
                   //Inner gross glass width [mm]
                   Chars_TO_Strg(Chars:=#AUX_rgcReceiveBuffer,
                                 pChars:=38,
                                 Cnt:=5,
                                 Strg=>#TMP_strValue);

                   #AUX_tYTelegram.dInLimitGross_mm := STRING_TO_DINT(#TMP_strValue); 

                   //Outer gross glass width [mm]
                   Chars_TO_Strg(Chars:=#AUX_rgcReceiveBuffer,
                                 pChars:=44,
                                 Cnt:=5,
                                 Strg=>#TMP_strValue);

                   #AUX_tYTelegram.dOutLimitGross_mm := STRING_TO_DINT(#TMP_strValue); 

                   //Center orientated position of the inner toproller [mm]
                   Chars_TO_Strg(Chars:=#AUX_rgcReceiveBuffer,
                                 pChars:=50,
                                 Cnt:=5,
                                 Strg=>#TMP_strValue);

                   #AUX_tYTelegram.dCenterOrientInTop_mm := STRING_TO_DINT(#TMP_strValue); 

                   //Edge orientated position of the inner toproller [mm]
                   Chars_TO_Strg(Chars:=#AUX_rgcReceiveBuffer,
                                 pChars:=56,
                                 Cnt:=5,
                                 Strg=>#TMP_strValue);

                   #AUX_tYTelegram.dEdgeOrientInTop_mm := STRING_TO_DINT(#TMP_strValue); 

                   //Center orientated position of the outer toproller [mm]
                   Chars_TO_Strg(Chars:=#AUX_rgcReceiveBuffer,
                                 pChars:=62,
                                 Cnt:=5,
                                 Strg=>#TMP_strValue);

                   #AUX_tYTelegram.dCenterOrientOutTop_mm := STRING_TO_DINT(#TMP_strValue); 

                   //Edge orientated position of the outer toproll [mm]
                   Chars_TO_Strg(Chars:=#AUX_rgcReceiveBuffer,
                                 pChars:=68,
                                 Cnt:=5,
                                 Strg=>#TMP_strValue);

                   #AUX_tYTelegram.dEdgeOrientOutTop_mm := STRING_TO_DINT(#TMP_strValue); 

                   //Check the conformity
                   IF #AUX_tYTelegram.dTelCounter < 0 OR
                      #AUX_tYTelegram.dTelCounter > 65535 OR
                      #AUX_tYTelegram.dFeedPulse_mm < 0 OR 
                      #AUX_tYTelegram.dFeedPulse_mm > 65535 OR
                      #AUX_tYTelegram.dInLimit_mm < 0 OR 
                      #AUX_tYTelegram.dInLimit_mm > 65535 OR
                      #AUX_tYTelegram.dOutLimit_mm < 0 OR 
                      #AUX_tYTelegram.dOutLimit_mm > 65535 OR
                      #AUX_tYTelegram.dInLimitUsable_mm < 0 OR 
                      #AUX_tYTelegram.dInLimitUsable_mm > 65535 OR
                      #AUX_tYTelegram.dOutLimitUsable_mm < 0 OR 
                      #AUX_tYTelegram.dOutLimitUsable_mm > 65535 OR
                      #AUX_tYTelegram.dInLimitGross_mm < 0 OR 
                      #AUX_tYTelegram.dInLimitGross_mm > 65535 OR
                      #AUX_tYTelegram.dOutLimitGross_mm < 0 OR 
                      #AUX_tYTelegram.dOutLimitGross_mm > 65535 OR
                      #AUX_tYTelegram.dCenterOrientInTop_mm < 0 OR 
                      #AUX_tYTelegram.dCenterOrientInTop_mm > 65535 OR
                      #AUX_tYTelegram.dEdgeOrientInTop_mm < 0 OR 
                      #AUX_tYTelegram.dEdgeOrientInTop_mm > 65535 OR
                      #AUX_tYTelegram.dCenterOrientOutTop_mm < 0 OR 
                      #AUX_tYTelegram.dCenterOrientOutTop_mm > 65535 OR
                      #AUX_tYTelegram.dEdgeOrientOutTop_mm < 0 OR 
                      #AUX_tYTelegram.dEdgeOrientOutTop_mm > 65535 THEN
                       #AUX_xTelegramYError := TRUE;
                   ELSE
                       IF #ST_xMachineSyncronized AND #tHMW.xAutoInspEnabled THEN

                           #TMP_dCountPos_cmm := #AUX_tYTelegram.dFeedPulse_mm - #AUX_dISRAValidCountMeter_mm;

                           IF #TMP_dCountPos_cmm < -32767 THEN

                               #AUX_tYTelegram.dPLCPosCount_cmm  := #AUX_dPLCValidCountMeter_cmm + ((#TMP_dCountPos_cmm + 65536)*100);

                           ELSIF #TMP_dCountPos_cmm > 32767 THEN

                               #AUX_tYTelegram.dPLCPosCount_cmm := #AUX_dPLCValidCountMeter_cmm + ((#TMP_dCountPos_cmm - 65536)*100);

                           ELSE

                               #AUX_tYTelegram.dPLCPosCount_cmm := #AUX_dPLCValidCountMeter_cmm + (#TMP_dCountPos_cmm * 100);

                           END_IF;

                           #AUX_tYTelegram.dPLCPosCount_cmm := #tHMR.dDistSnapRoll_cmm + #AUX_tYTelegram.dPLCPosCount_cmm;

                           #tHMR.dCurrentGrossWidth_cmm := (#AUX_tYTelegram.dOutLimitGross_mm - #AUX_tYTelegram.dInLimitGross_mm) * 100 ;
                           #tHMR.dCurrentNetWidth_cmm := (#AUX_tYTelegram.dOutLimitUsable_mm - #AUX_tYTelegram.dInLimitUsable_mm) * 100 ;

                           IF (#tHMR.dDistCenterLine_cmm <= 0) THEN

                               #tHMR.dCurrentGrossWander_cmm := #tHMR.dDistCenterLine_cmm + ((#AUX_tYTelegram.dInLimitGross_mm + #AUX_tYTelegram.dOutLimitGross_mm)/2) * 100;
                               #tHMR.dCurrentNetWander_cmm := #tHMR.dDistCenterLine_cmm + ((#AUX_tYTelegram.dInLimitUsable_mm + #AUX_tYTelegram.dOutLimitUsable_mm)/2) * 100;

                           ELSE
                               #tHMR.dCurrentGrossWander_cmm := #tHMR.dDistCenterLine_cmm - ((#AUX_tYTelegram.dInLimitGross_mm + #AUX_tYTelegram.dOutLimitGross_mm)/2) * 100;
                               #tHMR.dCurrentNetWander_cmm := #tHMR.dDistCenterLine_cmm - ((#AUX_tYTelegram.dInLimitUsable_mm + #AUX_tYTelegram.dOutLimitUsable_mm)/2) * 100;

                           END_IF;

                           #INO_tRibbon.rgtGlassData[#IN_dGlassDataMachineIndex].dDistSnapRoll_cmm := #tHMR.dDistSnapRoll_cmm + #DISRADEADPOINT_CMM; 

                           //Update the position
                           IF NOT #INO_tRibbon.rgtGlassDataUpdate[#IN_dGlassDataUpdateMachineIndex].xUpdateRequest THEN
                               #INO_tRibbon.rgtGlassDataUpdate[#IN_dGlassDataUpdateMachineIndex].tData.dGrossWander_cmm := #tHMR.dCurrentGrossWander_cmm;
                               #INO_tRibbon.rgtGlassDataUpdate[#IN_dGlassDataUpdateMachineIndex].tData.dNetWander_cmm := #tHMR.dCurrentNetWander_cmm;
                               #INO_tRibbon.rgtGlassDataUpdate[#IN_dGlassDataUpdateMachineIndex].tData.dGrossWidth_cmm := #tHMR.dCurrentGrossWidth_cmm;
                               #INO_tRibbon.rgtGlassDataUpdate[#IN_dGlassDataUpdateMachineIndex].tData.dNetWidth_cmm := #tHMR.dCurrentNetWidth_cmm;
                               #INO_tRibbon.rgtGlassDataUpdate[#IN_dGlassDataUpdateMachineIndex].xUpdateRequest := TRUE;
                           END_IF;
                       END_IF;
                   END_IF;
               END_IF;

             #DNUMCHAR_TEL_B_S:

               IF #AUX_rgcReceiveBuffer[0] = 'B' THEN


                   IF  #AUX_rgcReceiveBuffer[1] = ' ' AND
                       #AUX_rgcReceiveBuffer[7] = ' ' AND
                       #AUX_rgcReceiveBuffer[13] = #STR_CR AND
                       #AUX_rgcReceiveBuffer[14] = #STR_LF THEN

                        //Evaluate the data of the Y telegram
                       #TMP_dTelCount :=  #AUX_tBTelegram.dTelCounter;               

                       #TMP_dTelCount += 1;

                       IF #TMP_dTelCount >= 65535 THEN
                           #TMP_dTelCount := 1;
                       END_IF; 

                       Chars_TO_Strg(Chars:=#AUX_rgcReceiveBuffer,
                                     pChars:=2,
                                     Cnt:=5,
                                     Strg=>#TMP_strValue);

                       #AUX_tBTelegram.dTelCounter := STRING_TO_DINT(#TMP_strValue); 

                       IF (#TMP_dTelCount <> #AUX_tBTelegram.dTelCounter) THEN
                           #AUX_xTelegramBMissing := 1;    
                       END_IF;

                       Chars_TO_Strg(Chars:=#AUX_rgcReceiveBuffer,
                                     pChars:=8,
                                     Cnt:=5,
                                     Strg=>#TMP_strValue);

                       #AUX_tBTelegram.dFeedPulse_mm := STRING_TO_DINT(#TMP_strValue); 

                       //Check the conformity
                       IF  #AUX_tBTelegram.dTelCounter < 0 OR 
                           #AUX_tBTelegram.dTelCounter > 65535 OR
                           #AUX_tBTelegram.dFeedPulse_mm < 0 OR
                           #AUX_tBTelegram.dFeedPulse_mm > 65535 THEN                
                               #AUX_xTelegramBError := 1;  
                       ELSE
                           #AUX_tBTelegram.xNewTelegram := 1;
                       END_IF;
                   END_IF;
               ELSIF #AUX_rgcReceiveBuffer[0] = 'S' THEN

                   IF  #AUX_rgcReceiveBuffer[1] = ' ' AND
                       #AUX_rgcReceiveBuffer[7] = ' ' AND
                       #AUX_rgcReceiveBuffer[13] = #STR_CR AND
                       #AUX_rgcReceiveBuffer[14] = #STR_LF THEN

                        //Evaluate the data of the Y telegram
                       #TMP_dTelCount :=  #AUX_tSTelegram.dTelCounter;               

                       #TMP_dTelCount += 1;

                       IF #TMP_dTelCount >= 65535 THEN
                           #TMP_dTelCount := 1;
                       END_IF; 

                       Chars_TO_Strg(Chars:=#AUX_rgcReceiveBuffer,
                                     pChars:=2,
                                     Cnt:=5,
                                     Strg=>#TMP_strValue);

                       #AUX_tSTelegram.dTelCounter := STRING_TO_DINT(#TMP_strValue); 

                       IF (#TMP_dTelCount <> #AUX_tSTelegram.dTelCounter) THEN
                           #AUX_xTelegramSMissing := 1;    
                       END_IF;

                       Chars_TO_Strg(Chars:=#AUX_rgcReceiveBuffer,
                                     pChars:=8,
                                     Cnt:=5,
                                     Strg=>#TMP_strValue);

                       #AUX_tSTelegram.dFeedPulse_mm := STRING_TO_DINT(#TMP_strValue); 

                       //Check the conformity
                       IF  #AUX_tSTelegram.dTelCounter < 0 OR 
                           #AUX_tSTelegram.dTelCounter > 65535 OR
                           #AUX_tSTelegram.dFeedPulse_mm < 0 OR
                           #AUX_tSTelegram.dFeedPulse_mm > 65535 THEN                
                               #AUX_xTelegramSError := 1;  
                       ELSE
                           #AUX_tSTelegram.xNewTelegram := 1;
                       END_IF;
                   END_IF;

               ELSE
                   #AUX_xTelegramError := TRUE;             
               END_IF;            

           ELSE  // Statement section ELSE
               #AUX_xTelegramError := TRUE;
           END_CASE;

           //Take out the telegram read out and move up the buffer
           IF (#TMP_dCharCounter) < #AUX_dNumCharRecvBuffer THEN
               #TMP_iRetVal := MOVE_BLK_VARIANT(SRC:=#AUX_rgcReceiveBuffer, COUNT:=DINT_TO_UDINT(#AUX_dNumCharRecvBuffer - (#TMP_dCharCounter))   , SRC_INDEX:= #TMP_dCharCounter , DEST_INDEX:= 0, DEST=>#AUX_rgcReceiveBuffer);
               #AUX_dNumCharRecvBuffer -= #TMP_dCharCounter;
               #TMP_dCharCounter := 1;
               #TMP_dIndex := -1;
           ELSE
               #AUX_dNumCharRecvBuffer := 0;
           END_IF;
       END_IF;

       #TMP_dIndex+=1;

   END_WHILE;
END_REGION

REGION Network 20: Wait syncro data from scanner
   RUNG wire#powerrail
      Contact( #INO_tEncoder.xMeterForScanner )
      I_Contact( #tPh.xWaitSyncroData )
      wire#w1
      S_Coil( #tPh.xWaitSyncroData )
   END_RUNG
   RUNG wire#w1
      R_Coil( #INO_tEncoder.xMeterForScanner )
   END_RUNG
   // the same network as SCL:
   #_w1 := #INO_tEncoder.xMeterForScanner AND NOT #tPh.xWaitSyncroData;
   IF #_w1 THEN
       #tPh.xWaitSyncroData := TRUE;
       #INO_tEncoder.xMeterForScanner := FALSE;
   END_IF;
END_REGION

REGION Network 21: End wait syncro data from scanner
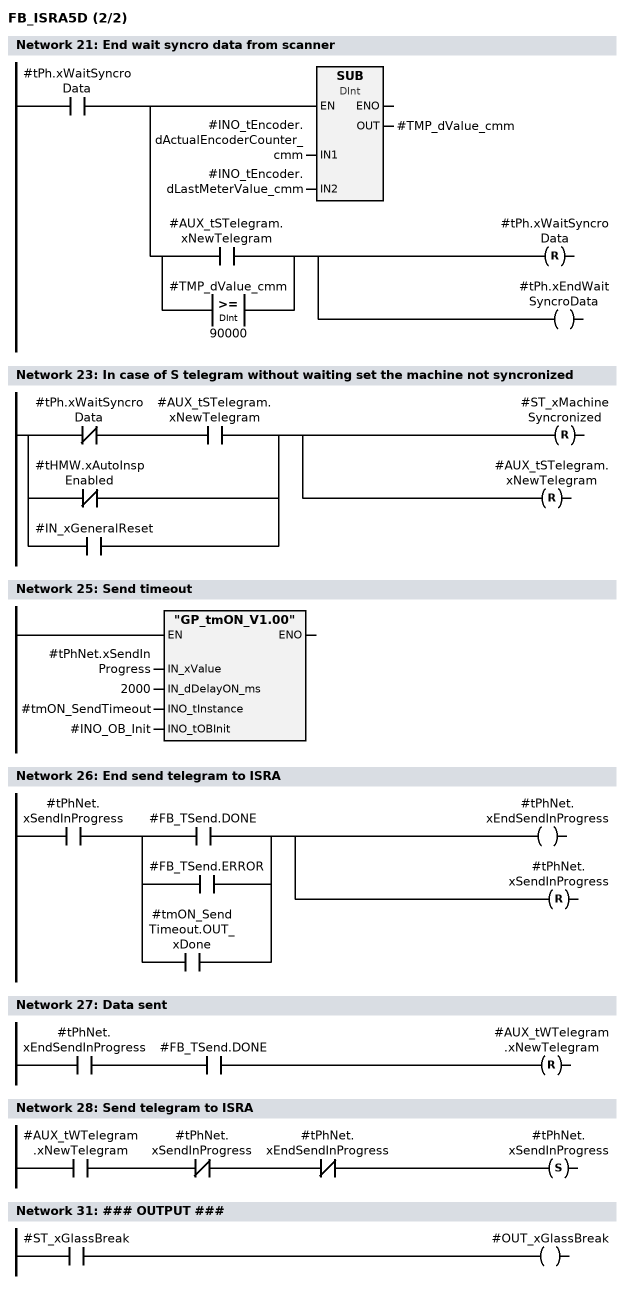
   RUNG wire#powerrail
      Contact( #tPh.xWaitSyncroData )
      wire#w1
      { S7_Templates := "SrcType := DInt" } Sub(in1 := #INO_tEncoder.dActualEncoderCounter_cmm, in2 := #INO_tEncoder.dLastMeterValue_cmm, out => #TMP_dValue_cmm)
   END_RUNG
   RUNG wire#w1
      Contact( #AUX_tSTelegram.xNewTelegram )
      wire#w2
      R_Coil( #tPh.xWaitSyncroData )
   END_RUNG
   RUNG wire#w1
      { S7_Templates := "SrcType := DInt" } GE_Contact(in1 := #TMP_dValue_cmm, in2 := 90000)
   END_RUNG wire#w2
   RUNG wire#w2
      Coil( #tPh.xEndWaitSyncroData )
   END_RUNG
   // the same network as SCL:
   IF #tPh.xWaitSyncroData THEN
       #TMP_dValue_cmm := #INO_tEncoder.dActualEncoderCounter_cmm - #INO_tEncoder.dLastMeterValue_cmm;
   END_IF;
   #_w1 := #tPh.xWaitSyncroData AND (#AUX_tSTelegram.xNewTelegram OR (#TMP_dValue_cmm >= 90000));
   IF #_w1 THEN #tPh.xWaitSyncroData := FALSE; END_IF;
   #tPh.xEndWaitSyncroData := #_w1;
END_REGION

REGION Network 22 (SCL): Set machine syncronized
   IF #tPh.xEndWaitSyncroData AND #AUX_tSTelegram.xNewTelegram THEN

       IF #ST_xMachineSyncronized THEN

           //This routine will validate if the syncro space is correct
           #TMP_dValue_cmm := #AUX_tSTelegram.dFeedPulse_mm - #AUX_dISRAValidCountMeter_mm;

           IF #TMP_dValue_cmm < -32767 THEN
               #TMP_dValue_cmm := #TMP_dValue_cmm + 65536;
           ELSIF #TMP_dValue_cmm > 32767 THEN
               #TMP_dValue_cmm := #TMP_dValue_cmm - 65536;
           END_IF;

           IF #TMP_dValue_cmm < 1100 AND #TMP_dValue_cmm > 900 THEN
               #AUX_dISRAValidCountMeter_mm := #AUX_tSTelegram.dFeedPulse_mm;
               #AUX_dPLCValidCountMeter_cmm := #INO_tEncoder.dLastMeterValue_cmm;
           ELSE
               #ST_xMachineSyncronized := FALSE;
               #OS_xSyncroOutLimits := TRUE; 
           END_IF;

       ELSE

           #AUX_dISRAValidCountMeter_mm := #AUX_tSTelegram.dFeedPulse_mm;
           #AUX_dPLCValidCountMeter_cmm := #INO_tEncoder.dLastMeterValue_cmm;
           #ST_xMachineSyncronized := TRUE;

       END_IF;

       #AUX_tSTelegram.xNewTelegram := FALSE;

   ELSIF #tPh.xEndWaitSyncroData AND NOT #AUX_tSTelegram.xNewTelegram THEN

       #ST_xMachineSyncronized := FALSE;
       #OS_xSyncroTimeout := TRUE;

   END_IF;
END_REGION

REGION Network 23: In case of S telegram without waiting set the machine not syncronized
   RUNG wire#powerrail
      I_Contact( #tPh.xWaitSyncroData )
      Contact( #AUX_tSTelegram.xNewTelegram )
      wire#w1
      R_Coil( #ST_xMachineSyncronized )
   END_RUNG
   RUNG wire#powerrail
      I_Contact( #tHMW.xAutoInspEnabled )
   END_RUNG wire#w1
   RUNG wire#powerrail
      Contact( #IN_xGeneralReset )
   END_RUNG wire#w1
   RUNG wire#w1
      R_Coil( #AUX_tSTelegram.xNewTelegram )
   END_RUNG
   // the same network as SCL:
   IF (NOT #tPh.xWaitSyncroData AND #AUX_tSTelegram.xNewTelegram) OR NOT #tHMW.xAutoInspEnabled OR #IN_xGeneralReset THEN
       #ST_xMachineSyncronized := FALSE;
       #AUX_tSTelegram.xNewTelegram := FALSE;
   END_IF;
END_REGION

REGION Network 24 (SCL): Prepare T telegram
   IF #AUX_tBTelegram.xNewTelegram THEN

       #AUX_tBTelegram.xNewTelegram := 0;

       //Increase the counter of telegram
       #AUX_tWTelegram.dTelCounter := #AUX_tWTelegram.dTelCounter + 1;

       IF #AUX_tWTelegram.dTelCounter > 65535 THEN
           #AUX_tWTelegram.dTelCounter := 0;
       END_IF;

       //The pulse counter is on decision line
       #AUX_tWTelegram.dFeedPulse_mm := #AUX_dISRAValidCountMeter_mm - ((#tHMR.dDistSnapRoll_cmm - #INO_tOptManager.tHMR.dDecisionLinePosition_cmm) / 100);

       IF (#AUX_tWTelegram.dFeedPulse_mm < 0) THEN
           #AUX_tWTelegram.dFeedPulse_mm := 65535 - #AUX_tWTelegram.dFeedPulse_mm; 
       END_IF;

       //Calculate the position
       #AUX_tWTelegram.dCutToolOpSide_mm := ((#INO_tCaps.tLastPlacedCap.dWidth_cmm / -2) +   #INO_tCaps.tLastPlacedCap.dEndCutWander_cmm)/ 100;

       //Normalize the value
       #AUX_tWTelegram.dCutToolOpSide_mm := ABS(#tHMR.dDistCenterLine_cmm / 100) + #AUX_tWTelegram.dCutToolOpSide_mm;

       #AUX_tWTelegram.dCutToolOppoOpSide_mm := #AUX_tWTelegram.dCutToolOpSide_mm + (#INO_tCaps.tLastPlacedCap.dWidth_cmm / 100);

       //Prepare the string to send
       //Fill to '0' the chars
       FOR #TMP_dIndex := 0 TO #DNUMCHAR_TEL_W_INDEX DO
           #AUX_rgsWTelegram[#TMP_dIndex] := '0'; //0
       END_FOR;


       #AUX_rgsWTelegram[0] := 'W'; //T
       #AUX_rgsWTelegram[1] := ' '; //Space

       #TMP_strValue := DINT_TO_STRING(#AUX_tWTelegram.dTelCounter);
       //Remove the sign
       #TMP_strValue := DELETE(IN:=#TMP_strValue, L:=1, P:=1);
       //Check the length
       #TMP_iStrLength := LEN(#TMP_strValue);
       //Move to the array
       Strg_TO_Chars(Strg:=#TMP_strValue,
                     pChars:=7 - #TMP_iStrLength,
                     Cnt=>#TMP_uiMovedChar,
                     Chars:=#AUX_rgsWTelegram);

       #AUX_rgsWTelegram[7] := ' '; //Space

       #TMP_strValue := DINT_TO_STRING(#AUX_tWTelegram.dFeedPulse_mm);
       //Remove the sign
       #TMP_strValue := DELETE(IN:=#TMP_strValue, L:=1, P:=1);
       //Check the length
       #TMP_iStrLength := LEN(#TMP_strValue);
       //Move to the array
       Strg_TO_Chars(Strg:=#TMP_strValue,
                     pChars:=13 - #TMP_iStrLength,
                     Cnt=>#TMP_uiMovedChar,
                     Chars:=#AUX_rgsWTelegram);

       #AUX_rgsWTelegram[13] := ' '; //Space

       #TMP_strValue := DINT_TO_STRING(#AUX_tWTelegram.dCutToolOpSide_mm + 100);
       //Remove the sign
       #TMP_strValue := DELETE(IN:=#TMP_strValue, L:=1, P:=1);
       //Check the length
       #TMP_iStrLength := LEN(#TMP_strValue);
       //Move to the array
       Strg_TO_Chars(Strg:=#TMP_strValue,
                     pChars:=19 - #TMP_iStrLength,
                     Cnt=>#TMP_uiMovedChar,
                     Chars:=#AUX_rgsWTelegram);

       #AUX_rgsWTelegram[19] := ' ' ; //Space

       #TMP_strValue := DINT_TO_STRING(#AUX_tWTelegram.dCutToolOppoOpSide_mm);
       //Remove the sign
       #TMP_strValue := DELETE(IN:=#TMP_strValue, L:=1, P:=1);
       //Check the length
       #TMP_iStrLength := LEN(#TMP_strValue);
       //Move to the array
       Strg_TO_Chars(Strg:=#TMP_strValue,
                     pChars:=25 - #TMP_iStrLength,
                     Cnt=>#TMP_uiMovedChar,
                     Chars:=#AUX_rgsWTelegram);

       #AUX_rgsWTelegram[25] := ' ' ; //Space

       #TMP_strValue := DINT_TO_STRING(#AUX_tWTelegram.dCutToolOpSide_mm);
       //Remove the sign
       #TMP_strValue := DELETE(IN:=#TMP_strValue, L:=1, P:=1);
       //Check the length
       #TMP_iStrLength := LEN(#TMP_strValue);
       //Move to the array
       Strg_TO_Chars(Strg:=#TMP_strValue,
                     pChars:=31 - #TMP_iStrLength,
                     Cnt=>#TMP_uiMovedChar,
                     Chars:=#AUX_rgsWTelegram);

       #AUX_rgsWTelegram[31] := ' ' ; //Space

       #TMP_strValue := DINT_TO_STRING(#AUX_tWTelegram.dCutToolOppoOpSide_mm);
       //Remove the sign
       #TMP_strValue := DELETE(IN:=#TMP_strValue, L:=1, P:=1);
       //Check the length
       #TMP_iStrLength := LEN(#TMP_strValue);
       //Move to the array
       Strg_TO_Chars(Strg:=#TMP_strValue,
                     pChars:=37 - #TMP_iStrLength,
                     Cnt=>#TMP_uiMovedChar,
                     Chars:=#AUX_rgsWTelegram);

       #AUX_rgsWTelegram[37] := #STR_CR; //CR
       #AUX_rgsWTelegram[38] := #STR_LF; //LF

       #AUX_tWTelegram.xNewTelegram := TRUE;
   END_IF;
END_REGION

REGION Network 25: Send timeout
   RUNG wire#powerrail
      "GP_tmON_V1.00"(IN_xValue := #tPhNet.xSendInProgress, IN_dDelayON_ms := 2000, INO_tInstance := #tmON_SendTimeout, INO_tOBInit := #INO_OB_Init)
   END_RUNG
   // the same network as SCL:
   "GP_tmON_V1.00"(IN_xValue := #tPhNet.xSendInProgress,
                   IN_dDelayON_ms := 2000,
                   INO_tInstance := #tmON_SendTimeout,
                   INO_tOBInit := #INO_OB_Init);
END_REGION

REGION Network 26: End send telegram to ISRA
   RUNG wire#powerrail
      Contact( #tPhNet.xSendInProgress )
      wire#w1
      Contact( #FB_TSend.DONE )
      wire#w2
      Coil( #tPhNet.xEndSendInProgress )
   END_RUNG
   RUNG wire#w1
      Contact( #FB_TSend.ERROR )
   END_RUNG wire#w2
   RUNG wire#w1
      Contact( #tmON_SendTimeout.OUT_xDone )
   END_RUNG wire#w2
   RUNG wire#w2
      R_Coil( #tPhNet.xSendInProgress )
   END_RUNG
   // the same network as SCL:
   #tPhNet.xEndSendInProgress := #tPhNet.xSendInProgress AND (#FB_TSend.DONE OR #FB_TSend.ERROR OR #tmON_SendTimeout.OUT_xDone);
   IF #tPhNet.xEndSendInProgress THEN #tPhNet.xSendInProgress := FALSE; END_IF;
END_REGION

REGION Network 27: Data sent
   RUNG wire#powerrail
      Contact( #tPhNet.xEndSendInProgress )
      Contact( #FB_TSend.DONE )
      R_Coil( #AUX_tWTelegram.xNewTelegram )
   END_RUNG
   // the same network as SCL:
   IF #tPhNet.xEndSendInProgress AND #FB_TSend.DONE THEN #AUX_tWTelegram.xNewTelegram := FALSE; END_IF;
END_REGION

REGION Network 28: Send telegram to ISRA
   RUNG wire#powerrail
      Contact( #AUX_tWTelegram.xNewTelegram )
      I_Contact( #tPhNet.xSendInProgress )
      I_Contact( #tPhNet.xEndSendInProgress )
      S_Coil( #tPhNet.xSendInProgress )
   END_RUNG
   // the same network as SCL:
   IF #AUX_tWTelegram.xNewTelegram AND NOT #tPhNet.xSendInProgress AND NOT #tPhNet.xEndSendInProgress THEN
       #tPhNet.xSendInProgress := TRUE;
   END_IF;
END_REGION

REGION Network 29 (SCL): Retrieve glass break
   #INO_tRibbon.rgtGlassBreakRequest[#IN_dGlassBreakIndexGet].IN_dDistanceSnaproll_cmm := #tHMR.dDistSnapRoll_cmm + #DISRADEADPOINT_CMM;
   #INO_tRibbon.rgtGlassBreakRequest[#IN_dGlassBreakIndexGet].IN_dDownstreamOffset_cmm := #CONST_DBREAKDOWNOFF_CMM;
   #INO_tRibbon.rgtGlassBreakRequest[#IN_dGlassBreakIndexGet].IN_dUpstreamOffset_cmm := #CONST_DBREAKUPOFF_CMM;

   IF #INO_tRibbon.rgtGlassBreakRequest[#IN_dGlassBreakIndexGet].OUT_xDataReady THEN
       #ST_xGlassBreak := #INO_tRibbon.rgtGlassBreakRequest[#IN_dGlassBreakIndexGet].OUT_xGlassBreak;
   END_IF;

   IF #INO_tRibbon.rgtGlassBreakRequest[#IN_dGlassBreakIndexGet].OUT_xDataReady OR NOT #INO_tRibbon.rgtGlassBreakRequest[#IN_dGlassBreakIndexGet].IN_xRequestGlassBreak THEN
       #INO_tRibbon.rgtGlassBreakRequest[#IN_dGlassBreakIndexGet].OUT_xDataReady := FALSE;
       #INO_tRibbon.rgtGlassBreakRequest[#IN_dGlassBreakIndexGet].IN_xRequestGlassBreak := TRUE;
   END_IF;
END_REGION

REGION Network 30 (SCL): ### HMI STATUS ###
   IF NOT #tHMW.xAutoInspEnabled THEN
       #tHMR.dInspectionStatus := 1;
   ELSIF #ST_xStoppedFaults THEN
       #tHMR.dInspectionStatus := 7;
   ELSE
       #tHMR.dInspectionStatus := 3;
   END_IF;

   IF #IN_xScannerON THEN
       #tHMR.xScannerON := true    ;
   ELSE
       #tHMR.xScannerON := False;
   END_IF;
END_REGION

REGION Network 31: ### OUTPUT ###
   RUNG wire#powerrail
      Contact( #ST_xGlassBreak )
      Coil( #OUT_xGlassBreak )
   END_RUNG
   // the same network as SCL:
   #OUT_xGlassBreak := #ST_xGlassBreak;
END_REGION

REGION Network 32 (SCL): ### SIMULATION ACTIVE ###
   IF #IN_xSimulationActive THEN

       IF (((#AUX_xSimDecModeGWidth) AND (#AUX_xSimIncModeGWidth)) OR ((NOT #AUX_xSimDecModeGWidth) AND (NOT #AUX_xSimIncModeGWidth))) THEN
           #AUX_xSimDecModeGWidth := TRUE;
           #AUX_xSimIncModeGWidth := FALSE;
       END_IF;

       IF (((#AUX_xSimDecModeNWidth) AND (#AUX_xSimIncModeNWidth)) OR ((NOT #AUX_xSimDecModeNWidth) AND (NOT #AUX_xSimIncModeNWidth))) THEN
           #AUX_xSimDecModeNWidth := TRUE;
           #AUX_xSimIncModeNWidth := FALSE;
       END_IF;

       IF (((#AUX_xSimDecModeWander) AND (#AUX_xSimIncModeWander)) OR ((NOT #AUX_xSimDecModeWander) AND (NOT #AUX_xSimIncModeWander))) THEN
           #AUX_xSimDecModeWander := TRUE;
           #AUX_xSimIncModeWander := FALSE;
       END_IF;

       IF (#AUX_xSimDecModeGWidth) THEN
           #AUX_dSimGrossWidth_cmm -= 1;
       ELSE
           #AUX_dSimGrossWidth_cmm += 1;
       END_IF;

       IF (#AUX_xSimDecModeNWidth) THEN
           #AUX_dSimNetWidth_cmm -= 1;
       ELSE
           #AUX_dSimNetWidth_cmm += 1;
       END_IF;

       IF (#AUX_xSimDecModeWander) THEN
           #AUX_dSimWander_cmm -= 1;
       ELSE
           #AUX_dSimWander_cmm += 1;
       END_IF;

       IF (#AUX_dSimGrossWidth_cmm < #DSIM_MINGROSSWIDTH_CMM) THEN 
           #AUX_xSimDecModeGWidth := FALSE;
           #AUX_xSimIncModeGWidth := TRUE;
       END_IF;

       IF (#AUX_dSimGrossWidth_cmm > #DSIM_MAXGROSSWIDTH_CMM) THEN
           #AUX_xSimDecModeGWidth := TRUE;
           #AUX_xSimIncModeGWidth := FALSE;
       END_IF;

       IF (#AUX_dSimNetWidth_cmm < #DSIM_MINNETWIDTH_CMM) THEN
           #AUX_xSimDecModeNWidth := FALSE;
           #AUX_xSimIncModeNWidth := TRUE;
       END_IF;

       IF (#AUX_dSimNetWidth_cmm > #DSIM_MAXNETWIDTH_CMM) THEN
           #AUX_xSimDecModeNWidth := TRUE;
           #AUX_xSimIncModeNWidth := FALSE;
       END_IF;

       IF (#AUX_dSimWander_cmm < #DSIM_MINNETWANDER_CMM) THEN
           #AUX_xSimDecModeWander := FALSE;
           #AUX_xSimIncModeWander := TRUE;
       END_IF;

       IF (#AUX_dSimWander_cmm > #DSIM_MAXNETWANDER_CMM) THEN
           #AUX_xSimDecModeWander := TRUE;
           #AUX_xSimIncModeWander := FALSE;
       END_IF;

       #INO_tRibbon.rgtGlassData[#IN_dGlassDataMachineIndex].dDistSnapRoll_cmm := #tHMR.dDistSnapRoll_cmm + #DISRADEADPOINT_CMM;

       #tHMR.dCurrentGrossWander_cmm := #AUX_dSimWander_cmm;
       #tHMR.dCurrentNetWander_cmm := #AUX_dSimWander_cmm;
       #tHMR.dCurrentGrossWidth_cmm := #AUX_dSimGrossWidth_cmm;
       #tHMR.dCurrentNetWidth_cmm := #AUX_dSimNetWidth_cmm;

       //Update the position
       IF (NOT #INO_tRibbon.rgtGlassDataUpdate[#IN_dGlassDataUpdateMachineIndex].xUpdateRequest) AND #INO_OB_Init.OUT_xOs_5s THEN

           #INO_tRibbon.rgtGlassDataUpdate[#IN_dGlassDataUpdateMachineIndex].tData.dGrossWander_cmm := #tHMR.dCurrentGrossWander_cmm;
           #INO_tRibbon.rgtGlassDataUpdate[#IN_dGlassDataUpdateMachineIndex].tData.dNetWander_cmm := #tHMR.dCurrentNetWander_cmm;
           #INO_tRibbon.rgtGlassDataUpdate[#IN_dGlassDataUpdateMachineIndex].tData.dGrossWidth_cmm := #tHMR.dCurrentGrossWidth_cmm;
           #INO_tRibbon.rgtGlassDataUpdate[#IN_dGlassDataUpdateMachineIndex].tData.dNetWidth_cmm := #tHMR.dCurrentNetWidth_cmm;
           #INO_tRibbon.rgtGlassDataUpdate[#IN_dGlassDataUpdateMachineIndex].xUpdateRequest := TRUE;

       END_IF;

   END_IF;
END_REGION
END_FUNCTION_BLOCK

FUNCTION_BLOCK "FB_ISRASNAP_V1.00"   // FB34, LAD
TITLE = Snaproll machine V1.00
{ S7_Optimized_Access := 'TRUE' }
VERSION : 0.1
   VAR_INPUT
      IN_dMachineIndex : DInt;   // Tracking machine index
      IN_xCycleON : Bool;   // Cycle ON
      IN_xGeneralReset : Bool;   // General reset
      IN_xResetAlarms : Bool;   // Reset alarms
      IN_xFaultsEnabled : Bool;   // Faults enabled
   END_VAR
   VAR_OUTPUT
      tOutputs : Struct   // Outputs
         xSnap : Bool;   // Snap signal
         xSnapQlt : Bool;   // Snap QLT
      END_STRUCT;
   END_VAR
   VAR_IN_OUT
      INO_tTrack : "UDT_CapData_Tracking";   // Tracking plate
      INO_tEnc : "UDT_Encoder";   // Encoder data
      INO_tObInit : "GP_OB_Initialize";   // OB initialize
   END_VAR
   VAR
      ST_xPhaseInProgress : Bool;   // Phases are in progress
      AUX_xValidUpCap : Bool;   // Upstream cap is valid
      AUX_xValidDwCap : Bool;   // Downstream cap is valid
      AUX_dUpCapIndex : DInt;   // Index of the upstream cap
      AUX_dDwCapIndex : DInt;   // Index of the downstream cap
      OS_xNewCapUp : Bool;   // New cap arrived upstream
      OS_xNewCapDw : Bool;   // New cap arrived downstream
      OS_xNewCap : Bool;   // New cap arrived
      AUX_xUpIsQuality : Bool;   // Upstream cap is a quality cap
      AUX_xDwIsQuality : Bool;   // Downstream cap is a quality cap
      tmONOFF_SnapSignal : "UDT_IECTONTOFF_V1.00";   // Time ON snap signal
      tmOFF_QltSignal : "UDT_IECTOFF_V1.00";   // Time OFF qlt signal
   END_VAR
   VAR CONSTANT
      DQLT_SNAP_REACT_MS : DInt := 50;   // Quality snap reaction time [ms]
      DSNAP_RETAIN_MS : DInt := 400;   // Snap retention time [ms]
   END_VAR
BEGIN

REGION Network 1: ####_CONSTANTS_####
END_REGION

REGION Network 2: ####_MATCH_####
END_REGION

REGION Network 3 (SCL): Move data information to tracking
   #INO_tTrack.rgtTrackMachine[#IN_dMachineIndex].tUserData.dSetDistanceSnap_cmm := 0;
   #INO_tTrack.rgtTrackMachine[#IN_dMachineIndex].tUserData.dSetMachReacTime_ms := #DQLT_SNAP_REACT_MS;
END_REGION

REGION Network 4 (SCL): Manage tracking call

   #OS_xNewCapUp := FALSE;
   #OS_xNewCapDw := FALSE;
   #OS_xNewCap := FALSE;

   IF #INO_tTrack.rgtTrackMachine[#IN_dMachineIndex].tUserData.xGetPosReach THEN

       IF (NOT #ST_xPhaseInProgress) THEN

           #OS_xNewCap := TRUE;

           IF #INO_tTrack.rgtTrackMachine[#IN_dMachineIndex].tUserData.dGetUpstremIndex >= 0 THEN
               #AUX_xValidUpCap := TRUE;
               #OS_xNewCapUp := TRUE;            
               #AUX_dUpCapIndex := #INO_tTrack.rgtTrackMachine[#IN_dMachineIndex].tUserData.dGetUpstremIndex;

               IF  #INO_tTrack.rgtTrackCaps[#AUX_dUpCapIndex].tCap.rgtLites[0].dMainDestination = "DQUALITYDESTMASK1" OR
                   #INO_tTrack.rgtTrackCaps[#AUX_dUpCapIndex].tCap.rgtLites[0].dMainDestination = "DQUALITYDESTMASK2" OR
                   #INO_tTrack.rgtTrackCaps[#AUX_dUpCapIndex].tCap.rgtLites[0].dMainDestination = "DQUALITYDESTMASK3" OR
                   #INO_tTrack.rgtTrackCaps[#AUX_dUpCapIndex].tCap.rgtLites[0].dMainDestination = "DQUALITYDESTMASK4"
               THEN

                   #AUX_xUpIsQuality := TRUE;

               ELSE

                   #AUX_xUpIsQuality := FALSE;

               END_IF;

           ELSE
               #AUX_xValidUpCap := FALSE;
               #OS_xNewCapUp := FALSE;            
               #AUX_dUpCapIndex := 0;
           END_IF;

           IF #INO_tTrack.rgtTrackMachine[#IN_dMachineIndex].tUserData.dGetDownstreamIndex >= 0 THEN
               #AUX_xValidDwCap := TRUE;
               #OS_xNewCapDw := TRUE;            
               #AUX_dDwCapIndex := #INO_tTrack.rgtTrackMachine[#IN_dMachineIndex].tUserData.dGetDownstreamIndex;
           ELSE
               #AUX_xValidDwCap := FALSE;
               #OS_xNewCapDw := FALSE;            
               #AUX_dDwCapIndex := 0;
           END_IF;



       END_IF;

       #INO_tTrack.rgtTrackMachine[#IN_dMachineIndex].tUserData.xGetPosReach := FALSE;

   END_IF;
END_REGION

REGION Network 5: ####_HMI_LOGICS_####
END_REGION

REGION Network 6: ####_PHASES_&_LOGICS_####
END_REGION

REGION Network 7: Qlt Signal
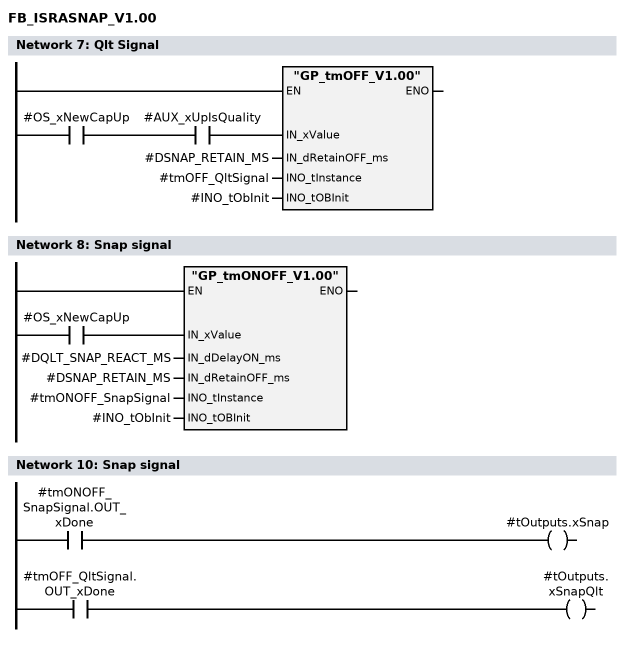
   RUNG wire#powerrail
      "GP_tmOFF_V1.00"(IN_xValue := wire#w1, IN_dRetainOFF_ms := #DSNAP_RETAIN_MS, INO_tInstance := #tmOFF_QltSignal, INO_tOBInit := #INO_tObInit)
   END_RUNG
   RUNG wire#powerrail
      Contact( #OS_xNewCapUp )
      Contact( #AUX_xUpIsQuality )
   END_RUNG wire#w1
   // the same network as SCL:
   "GP_tmOFF_V1.00"(IN_xValue := #OS_xNewCapUp AND #AUX_xUpIsQuality,
                    IN_dRetainOFF_ms := #DSNAP_RETAIN_MS,
                    INO_tInstance := #tmOFF_QltSignal,
                    INO_tOBInit := #INO_tObInit);
END_REGION

REGION Network 8: Snap signal
   RUNG wire#powerrail
      "GP_tmONOFF_V1.00"(IN_xValue := wire#w1, IN_dDelayON_ms := #DQLT_SNAP_REACT_MS, IN_dRetainOFF_ms := #DSNAP_RETAIN_MS, INO_tInstance := #tmONOFF_SnapSignal, INO_tOBInit := #INO_tObInit)
   END_RUNG
   RUNG wire#powerrail
      Contact( #OS_xNewCapUp )
   END_RUNG wire#w1
   // the same network as SCL:
   "GP_tmONOFF_V1.00"(IN_xValue := #OS_xNewCapUp,
                      IN_dDelayON_ms := #DQLT_SNAP_REACT_MS,
                      IN_dRetainOFF_ms := #DSNAP_RETAIN_MS,
                      INO_tInstance := #tmONOFF_SnapSignal,
                      INO_tOBInit := #INO_tObInit);
END_REGION

REGION Network 9: ####_OUTPUT_####
END_REGION

REGION Network 10: Snap signal
   RUNG wire#powerrail
      Contact( #tmONOFF_SnapSignal.OUT_xDone )
      Coil( #tOutputs.xSnap )
   END_RUNG
   RUNG wire#powerrail
      Contact( #tmOFF_QltSignal.OUT_xDone )
      Coil( #tOutputs.xSnapQlt )
   END_RUNG
   // the same network as SCL:
   #tOutputs.xSnap := #tmONOFF_SnapSignal.OUT_xDone;
   #tOutputs.xSnapQlt := #tmOFF_QltSignal.OUT_xDone;
END_REGION
END_FUNCTION_BLOCK

// folder: 03_Programs_Logics/MCC1200/20_Oil

FUNCTION_BLOCK "FB_Oil_V1.00"   // FB25, LAD
{ S7_Optimized_Access := 'TRUE' }
VERSION : 0.1
   VAR_INPUT
      IN_xCycleON : Bool;   // Cycle ON
      IN_xCycleONDel : Bool;   // Delayed cycle ON signal
      IN_xGeneralReset : Bool;   // General reset
      IN_xResetAlarms : Bool;   // Reset alarms
      IN_xFaultsEnabled : Bool;   // Faults enabled
      INPUT : Struct   // Digital inputs
         xOilMinLevel : Bool;   // L.Tank oil min level
         xOilMaxLevel : Bool;   // L.Tank oil max level
         xPowerSupply : Bool;   // L+.Power supply control
      END_STRUCT;
   END_VAR
   VAR_OUTPUT
      OUTPUT : Struct
         xTankFillCut : Bool;   // Y.Tank filling cutting
      END_STRUCT;
   END_VAR
   VAR_IN_OUT
      INO_tOBInitialize : "GP_OB_Initialize";   // OB Initialize
   END_VAR
   VAR
      tHMW : Struct   // HMI Write
         tMan : Struct   // Manual commands
            xFillTank : Bool;   // Fill tank {x|x|x|x|O}
            xSpare_1 : Bool;
            xSpare_2 : Bool;
            xSpare_3 : Bool;
            xSpare_4 : Bool;
            xSpare_5 : Bool;
            xSpare_6 : Bool;
            xSpare_7 : Bool;
            xSpare_8 : Bool;
            xSpare_9 : Bool;
            xSpare_10 : Bool;
            xSpare_11 : Bool;
            xSpare_12 : Bool;
            xSpare_13 : Bool;
            xSpare_14 : Bool;
            xSpare_15 : Bool;
         END_STRUCT;
         xEnDisManCom : Bool;   // Enable disable manual command {x|x|x|x|O}
      END_STRUCT;
      tHMR : Struct   // HMI Read
         dStatus : DInt;   // Status (1=Idle 3=Run 7=Anomaly) {X|X|X|X|O}
         xOilAtMin : Bool;   // Oil at minimum {X|X|X|X|O}
         xOilAtMax : Bool;   // Oil at maximum {X|X|X|X|O}
         xManComEn : Bool;   // Manual command enabled {x|x|x|x|O}
         tManFdbk : Struct   // Manual commands feedback
            xFillTank : Bool;   // Fill tank {x|x|x|x|O}
            xSpare_1 : Bool;
            xSpare_2 : Bool;
            xSpare_3 : Bool;
            xSpare_4 : Bool;
            xSpare_5 : Bool;
            xSpare_6 : Bool;
            xSpare_7 : Bool;
            xSpare_8 : Bool;
            xSpare_9 : Bool;
            xSpare_10 : Bool;
            xSpare_11 : Bool;
            xSpare_12 : Bool;
            xSpare_13 : Bool;
            xSpare_14 : Bool;
            xSpare_15 : Bool;
         END_STRUCT;
      END_STRUCT;
      tALM : Struct   // HMI Alarms
         tS : Struct   // Stopping faults machine
            xPowerSupplyControl : Bool;   // L+.Power supply control {X|X|X|X|O}
            xOilMinimumLevel : Bool;   // SL1.Oil at minimum {X|X|X|X|O}
            xTimeoutRefillOil : Bool;   // SL2.Timeout refill oil {X|X|X|X|O}
            xSensorMismatch : Bool;   // SL1/2.Sensor mismatch {X|X|X|X|O}
            xSpare_4 : Bool;
            xSpare_5 : Bool;
            xSpare_6 : Bool;
            xSpare_7 : Bool;
            xSpare_8 : Bool;
            xSpare_9 : Bool;
            xSpare_10 : Bool;
            xSpare_11 : Bool;
            xSpare_12 : Bool;
            xSpare_13 : Bool;
            xSpare_14 : Bool;
            xSpare_15 : Bool;
            xSpare_16 : Bool;
            xSpare_17 : Bool;
            xSpare_18 : Bool;
            xSpare_19 : Bool;
            xSpare_20 : Bool;
            xSpare_21 : Bool;
            xSpare_22 : Bool;
            xSpare_23 : Bool;
            xSpare_24 : Bool;
            xSpare_25 : Bool;
            xSpare_26 : Bool;
            xSpare_27 : Bool;
            xSpare_28 : Bool;
            xSpare_29 : Bool;
            xSpare_30 : Bool;
            xSpare_31 : Bool;
         END_STRUCT;
         tF : Struct   // Faults
            xSpare_0 : Bool;
            xSpare_1 : Bool;
            xSpare_2 : Bool;
            xSpare_3 : Bool;
            xSpare_4 : Bool;
            xSpare_5 : Bool;
            xSpare_6 : Bool;
            xSpare_7 : Bool;
            xSpare_8 : Bool;
            xSpare_9 : Bool;
            xSpare_10 : Bool;
            xSpare_11 : Bool;
            xSpare_12 : Bool;
            xSpare_13 : Bool;
            xSpare_14 : Bool;
            xSpare_15 : Bool;
            xSpare_16 : Bool;
            xSpare_17 : Bool;
            xSpare_18 : Bool;
            xSpare_19 : Bool;
            xSpare_20 : Bool;
            xSpare_21 : Bool;
            xSpare_22 : Bool;
            xSpare_23 : Bool;
            xSpare_24 : Bool;
            xSpare_25 : Bool;
            xSpare_26 : Bool;
            xSpare_27 : Bool;
            xSpare_28 : Bool;
            xSpare_29 : Bool;
            xSpare_30 : Bool;
            xSpare_31 : Bool;
         END_STRUCT;
         tW : Struct   // Warnings
            xSpare_0 : Bool;
            xSpare_1 : Bool;
            xSpare_2 : Bool;
            xSpare_3 : Bool;
            xSpare_4 : Bool;
            xSpare_5 : Bool;
            xSpare_6 : Bool;
            xSpare_7 : Bool;
            xSpare_8 : Bool;
            xSpare_9 : Bool;
            xSpare_10 : Bool;
            xSpare_11 : Bool;
            xSpare_12 : Bool;
            xSpare_13 : Bool;
            xSpare_14 : Bool;
            xSpare_15 : Bool;
            xSpare_16 : Bool;
            xSpare_17 : Bool;
            xSpare_18 : Bool;
            xSpare_19 : Bool;
            xSpare_20 : Bool;
            xSpare_21 : Bool;
            xSpare_22 : Bool;
            xSpare_23 : Bool;
            xSpare_24 : Bool;
            xSpare_25 : Bool;
            xSpare_26 : Bool;
            xSpare_27 : Bool;
            xSpare_28 : Bool;
            xSpare_29 : Bool;
            xSpare_30 : Bool;
            xSpare_31 : Bool;
         END_STRUCT;
      END_STRUCT;
      ST_xOutputEnable : Bool;   // Output enable
      ST_xCondOkMan : Bool;   // Condition ok manual command
      ST_xStoppedFaults : Bool;   // Stopped faults
      ST_xFaults : Bool;   // Faults
      ST_xWarning : Bool;   // Warnings
      ST_xRefillReq : Bool;   // Refill request
      AUX_tmOn_OilAtMinimum : "UDT_IECTON_V1.00";   // Oil at minimum level
      AUX_tmOn_TimeoutRefill : "UDT_IECTON_V1.00";   // Refill timeout
   END_VAR
   VAR_TEMP
      TMP_dwValue : DWord;
   END_VAR
   VAR CONSTANT
      CONST_DSTATUS_ANOMALY : DInt := 7;
      CONST_DSTATUS_RUN : DInt := 3;
      CONST_DSTATUS_IDLE : DInt := 1;
      CONST_DTIMEOUT_MS : DInt := 400000;   // Refill timeout [ms]
   END_VAR
   VAR_TEMP   // added for the SCL form of the ladder/FBD networks
      _w1 : Bool;
   END_VAR
BEGIN

REGION Network 1: ####_CONSTANTS_####
END_REGION

REGION Network 2: ####_MATCH_####
END_REGION

REGION Network 3: ####_HMI_LOGICS_####
END_REGION

REGION Network 4: Manual command enabled
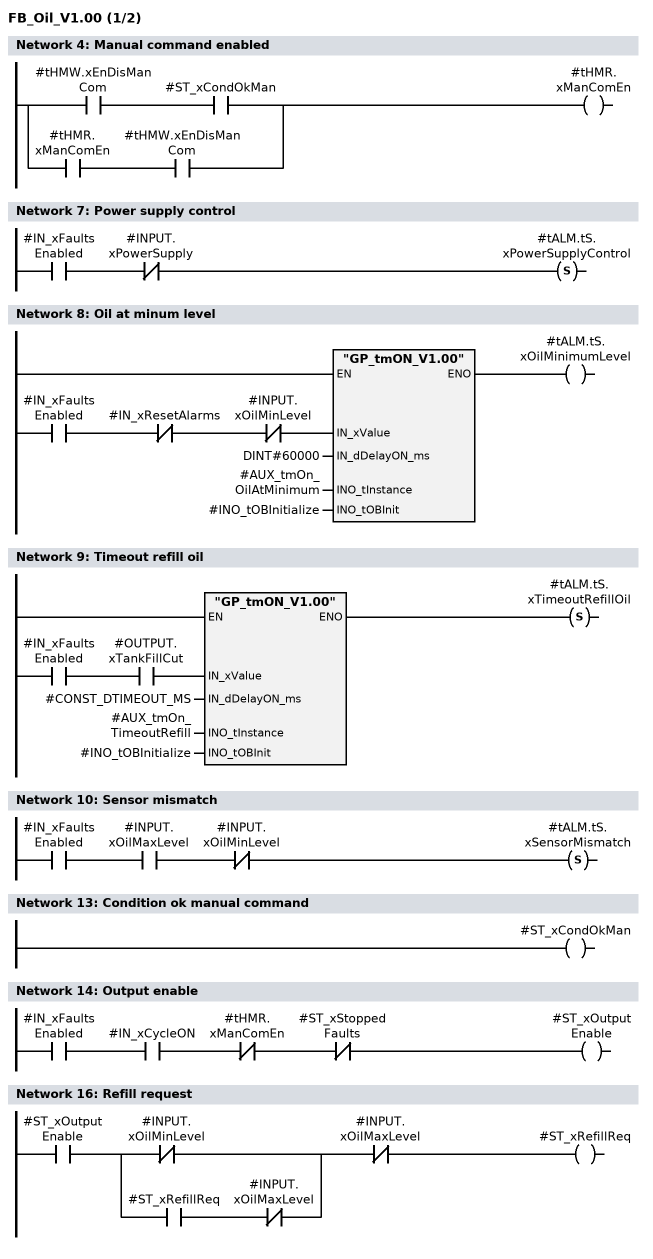
   RUNG wire#powerrail
      Contact( #tHMW.xEnDisManCom )
      Contact( #ST_xCondOkMan )
      wire#w1
      Coil( #tHMR.xManComEn )
   END_RUNG
   RUNG wire#powerrail
      Contact( #tHMR.xManComEn )
      Contact( #tHMW.xEnDisManCom )
   END_RUNG wire#w1
   // the same network as SCL:
   #tHMR.xManComEn := (#tHMW.xEnDisManCom AND #ST_xCondOkMan) OR (#tHMR.xManComEn AND #tHMW.xEnDisManCom);
END_REGION

REGION Network 5: ####_ALARMS_####
END_REGION

REGION Network 6 (SCL): Reset alarms
   IF #IN_xResetAlarms THEN

       #TMP_dwValue := 0;

       SCATTER(IN:=#TMP_dwValue,
               OUT=>#tALM.tS);

       SCATTER(IN:=#TMP_dwValue,
               OUT=>#tALM.tF);

       SCATTER(IN:=#TMP_dwValue,
               OUT=>#tALM.tW);


   END_IF;
END_REGION

REGION Network 7: Power supply control
   RUNG wire#powerrail
      Contact( #IN_xFaultsEnabled )
      I_Contact( #INPUT.xPowerSupply )
      S_Coil( #tALM.tS.xPowerSupplyControl )
   END_RUNG
   // the same network as SCL:
   IF #IN_xFaultsEnabled AND NOT #INPUT.xPowerSupply THEN #tALM.tS.xPowerSupplyControl := TRUE; END_IF;
END_REGION

REGION Network 8: Oil at minum level
   RUNG wire#powerrail
      "GP_tmON_V1.00"(IN_xValue := wire#w1, IN_dDelayON_ms := DINT#60000, INO_tInstance := #AUX_tmOn_OilAtMinimum, INO_tOBInit := #INO_tOBInitialize)
      Coil( #tALM.tS.xOilMinimumLevel )
   END_RUNG
   RUNG wire#powerrail
      Contact( #IN_xFaultsEnabled )
      I_Contact( #IN_xResetAlarms )
      I_Contact( #INPUT.xOilMinLevel )
   END_RUNG wire#w1
   // the same network as SCL:
   "GP_tmON_V1.00"(IN_xValue := #IN_xFaultsEnabled AND NOT #IN_xResetAlarms AND NOT #INPUT.xOilMinLevel,
                   IN_dDelayON_ms := DINT#60000,
                   INO_tInstance := #AUX_tmOn_OilAtMinimum,
                   INO_tOBInit := #INO_tOBInitialize,
                   ENO => #_w1);
   #tALM.tS.xOilMinimumLevel := #_w1;
END_REGION

REGION Network 9: Timeout refill oil
   RUNG wire#powerrail
      "GP_tmON_V1.00"(IN_xValue := wire#w1, IN_dDelayON_ms := #CONST_DTIMEOUT_MS, INO_tInstance := #AUX_tmOn_TimeoutRefill, INO_tOBInit := #INO_tOBInitialize)
      S_Coil( #tALM.tS.xTimeoutRefillOil )
   END_RUNG
   RUNG wire#powerrail
      Contact( #IN_xFaultsEnabled )
      Contact( #OUTPUT.xTankFillCut )
   END_RUNG wire#w1
   // the same network as SCL:
   "GP_tmON_V1.00"(IN_xValue := #IN_xFaultsEnabled AND #OUTPUT.xTankFillCut,
                   IN_dDelayON_ms := #CONST_DTIMEOUT_MS,
                   INO_tInstance := #AUX_tmOn_TimeoutRefill,
                   INO_tOBInit := #INO_tOBInitialize,
                   ENO => #_w1);
   IF #_w1 THEN #tALM.tS.xTimeoutRefillOil := TRUE; END_IF;
END_REGION

REGION Network 10: Sensor mismatch
   RUNG wire#powerrail
      Contact( #IN_xFaultsEnabled )
      Contact( #INPUT.xOilMaxLevel )
      I_Contact( #INPUT.xOilMinLevel )
      S_Coil( #tALM.tS.xSensorMismatch )
   END_RUNG
   // the same network as SCL:
   IF #IN_xFaultsEnabled AND #INPUT.xOilMaxLevel AND NOT #INPUT.xOilMinLevel THEN
       #tALM.tS.xSensorMismatch := TRUE;
   END_IF;
END_REGION

REGION Network 11 (SCL): Calculate comulative statuses
       GATHER(IN:=#tALM.tS,
              OUT=>#TMP_dwValue);

       IF #TMP_dwValue <> 0 THEN
           #ST_xStoppedFaults := TRUE;
       ELSE
           #ST_xStoppedFaults := FALSE;
       END_IF;

       GATHER(IN:=#tALM.tF,
              OUT=>#TMP_dwValue);

       IF #TMP_dwValue <> 0 THEN
           #ST_xFaults := TRUE;
       ELSE
           #ST_xFaults := FALSE;
       END_IF;

       GATHER(IN:=#tALM.tW,
              OUT=>#TMP_dwValue);

       IF #TMP_dwValue <> 0 THEN
           #ST_xWarning := TRUE;
       ELSE
           #ST_xWarning := FALSE;
       END_IF;
END_REGION

REGION Network 12: ####_STATUSES_####
END_REGION

REGION Network 13: Condition ok manual command
   RUNG wire#powerrail
      Coil( #ST_xCondOkMan )
   END_RUNG
   // the same network as SCL:
   #ST_xCondOkMan := TRUE;
END_REGION

REGION Network 14: Output enable
   RUNG wire#powerrail
      Contact( #IN_xFaultsEnabled )
      Contact( #IN_xCycleON )
      I_Contact( #tHMR.xManComEn )
      I_Contact( #ST_xStoppedFaults )
      Coil( #ST_xOutputEnable )
   END_RUNG
   // the same network as SCL:
   #ST_xOutputEnable := #IN_xFaultsEnabled AND #IN_xCycleON AND NOT #tHMR.xManComEn AND NOT #ST_xStoppedFaults;
END_REGION

REGION Network 15: ### PHASE AND LOGICS ###
END_REGION

REGION Network 16: Refill request
   RUNG wire#powerrail
      Contact( #ST_xOutputEnable )
      wire#w1
      I_Contact( #INPUT.xOilMinLevel )
      wire#w2
      I_Contact( #INPUT.xOilMaxLevel )
      Coil( #ST_xRefillReq )
   END_RUNG
   RUNG wire#w1
      Contact( #ST_xRefillReq )
      I_Contact( #INPUT.xOilMaxLevel )
   END_RUNG wire#w2
   // the same network as SCL:
   #ST_xRefillReq := #ST_xOutputEnable AND (NOT #INPUT.xOilMinLevel OR (#ST_xRefillReq AND NOT #INPUT.xOilMaxLevel)) AND NOT #INPUT.xOilMaxLevel;
END_REGION

REGION Network 17 (SCL): ### HMI STATUS ###
   IF #ST_xStoppedFaults THEN
       #tHMR.dStatus := #CONST_DSTATUS_ANOMALY;
   ELSIF #OUTPUT.xTankFillCut THEN
       #tHMR.dStatus := #CONST_DSTATUS_RUN;
   ELSE
       #tHMR.dStatus := #CONST_DSTATUS_IDLE;
   END_IF;

   #tHMR.xOilAtMin := #INPUT.xOilMinLevel;
   #tHMR.xOilAtMax := #INPUT.xOilMaxLevel;

   #tHMR.tManFdbk.xFillTank := #OUTPUT.xTankFillCut AND #tHMW.tMan.xFillTank;
END_REGION

REGION Network 18: ####_OUTPUT_####
END_REGION

REGION Network 19: Refill request
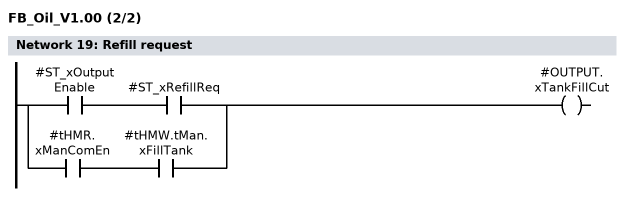
   RUNG wire#powerrail
      Contact( #ST_xOutputEnable )
      Contact( #ST_xRefillReq )
      wire#w1
      Coil( #OUTPUT.xTankFillCut )
   END_RUNG
   RUNG wire#powerrail
      Contact( #tHMR.xManComEn )
      Contact( #tHMW.tMan.xFillTank )
   END_RUNG wire#w1
   // the same network as SCL:
   #OUTPUT.xTankFillCut := (#ST_xOutputEnable AND #ST_xRefillReq) OR (#tHMR.xManComEn AND #tHMW.tMan.xFillTank);
END_REGION
END_FUNCTION_BLOCK

// folder: 03_Programs_Logics/MCC1200/21_Manual_Inspection

